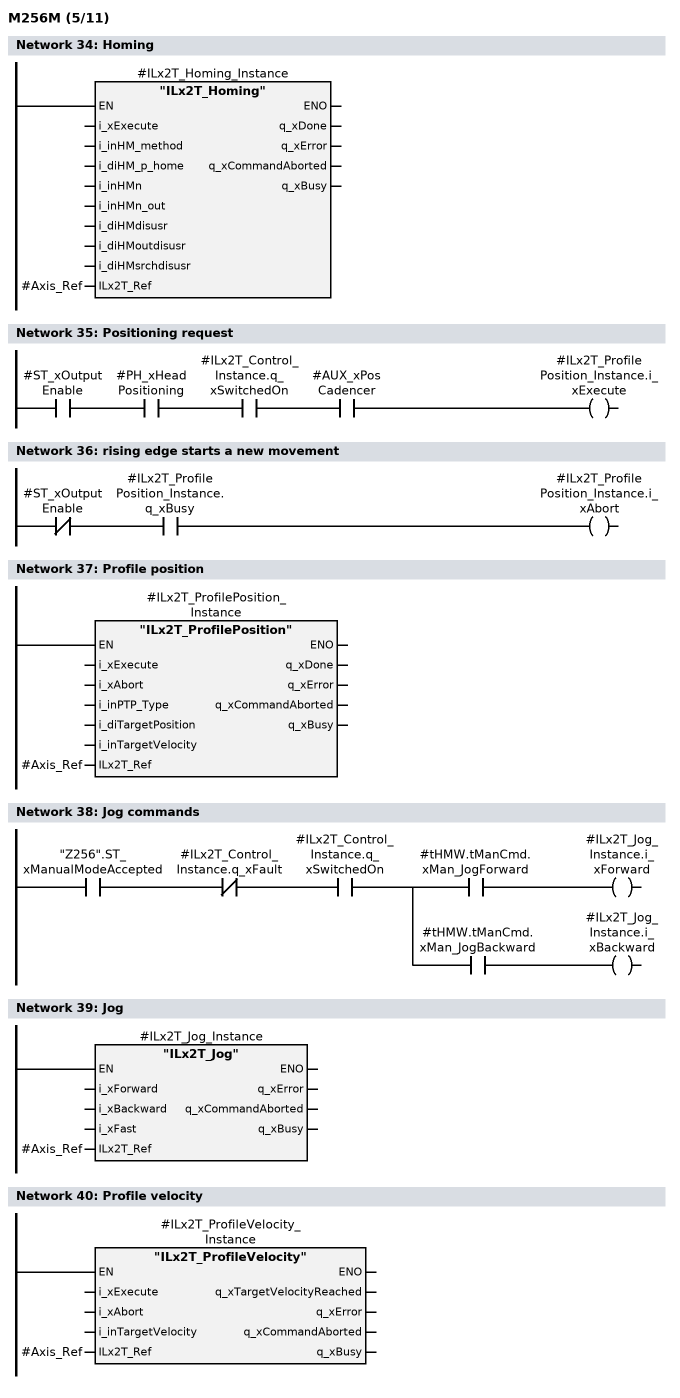
   RUNG wire#powerrail
      #ILx2T_Homing_Instance(i_xExecute :=, i_inHM_method :=, i_diHM_p_home :=, i_inHMn :=, i_inHMn_out :=, i_diHMdisusr :=, i_diHMoutdisusr :=, i_diHMsrchdisusr :=, ILx2T_Ref := #Axis_Ref, q_xDone =>, q_xError =>, q_xCommandAborted =>, q_xBusy =>)
   END_RUNG
   // the same network as SCL:
   #ILx2T_Homing_Instance(ILx2T_Ref := #Axis_Ref);   // "ILx2T_Homing"
END_REGION

REGION Network 35: Positioning request
   RUNG wire#powerrail
      Contact( #ST_xOutputEnable )
      Contact( #PH_xHeadPositioning )
      Contact( #ILx2T_Control_Instance.q_xSwitchedOn )
      Contact( #AUX_xPosCadencer )
      Coil( #ILx2T_ProfilePosition_Instance.i_xExecute )
   END_RUNG
   // the same network as SCL:
   #ILx2T_ProfilePosition_Instance.i_xExecute := #ST_xOutputEnable AND #PH_xHeadPositioning AND #ILx2T_Control_Instance.q_xSwitchedOn AND #AUX_xPosCadencer;
END_REGION

REGION Network 36: rising edge starts a new movement
   RUNG wire#powerrail
      I_Contact( #ST_xOutputEnable )
      Contact( #ILx2T_ProfilePosition_Instance.q_xBusy )
      Coil( #ILx2T_ProfilePosition_Instance.i_xAbort )
   END_RUNG
   // the same network as SCL:
   #ILx2T_ProfilePosition_Instance.i_xAbort := NOT #ST_xOutputEnable AND #ILx2T_ProfilePosition_Instance.q_xBusy;
END_REGION

REGION Network 37: Profile position
   RUNG wire#powerrail
      #ILx2T_ProfilePosition_Instance(i_xExecute :=, i_xAbort :=, i_inPTP_Type :=, i_diTargetPosition :=, i_inTargetVelocity :=, ILx2T_Ref := #Axis_Ref, q_xDone =>, q_xError =>, q_xCommandAborted =>, q_xBusy =>)
   END_RUNG
   // the same network as SCL:
   #ILx2T_ProfilePosition_Instance(ILx2T_Ref := #Axis_Ref);   // "ILx2T_ProfilePosition"
END_REGION

REGION Network 38: Jog commands
   RUNG wire#powerrail
      Contact( "Z256".ST_xManualModeAccepted )
      I_Contact( #ILx2T_Control_Instance.q_xFault )
      Contact( #ILx2T_Control_Instance.q_xSwitchedOn )
      wire#w1
      Contact( #tHMW.tManCmd.xMan_JogForward )
      Coil( #ILx2T_Jog_Instance.i_xForward )
   END_RUNG
   RUNG wire#w1
      Contact( #tHMW.tManCmd.xMan_JogBackward )
      Coil( #ILx2T_Jog_Instance.i_xBackward )
   END_RUNG
   // the same network as SCL:
   #_w1 := "Z256".ST_xManualModeAccepted AND NOT #ILx2T_Control_Instance.q_xFault AND #ILx2T_Control_Instance.q_xSwitchedOn;
   #ILx2T_Jog_Instance.i_xForward := #_w1 AND #tHMW.tManCmd.xMan_JogForward;
   #ILx2T_Jog_Instance.i_xBackward := #_w1 AND #tHMW.tManCmd.xMan_JogBackward;
END_REGION

REGION Network 39: Jog
   RUNG wire#powerrail
      #ILx2T_Jog_Instance(i_xForward :=, i_xBackward :=, i_xFast :=, ILx2T_Ref := #Axis_Ref, q_xError =>, q_xCommandAborted =>, q_xBusy =>)
   END_RUNG
   // the same network as SCL:
   #ILx2T_Jog_Instance(ILx2T_Ref := #Axis_Ref);   // "ILx2T_Jog"
END_REGION

REGION Network 40: Profile velocity
   RUNG wire#powerrail
      #ILx2T_ProfileVelocity_Instance(i_xExecute :=, i_xAbort :=, i_inTargetVelocity :=, ILx2T_Ref := #Axis_Ref, q_xTargetVelocityReached =>, q_xError =>, q_xCommandAborted =>, q_xBusy =>)
   END_RUNG
   // the same network as SCL:
   #ILx2T_ProfileVelocity_Instance(ILx2T_Ref := #Axis_Ref);   // "ILx2T_ProfileVelocity"
END_REGION

REGION Network 41: Head brake release
   // state 3=switch on disabled
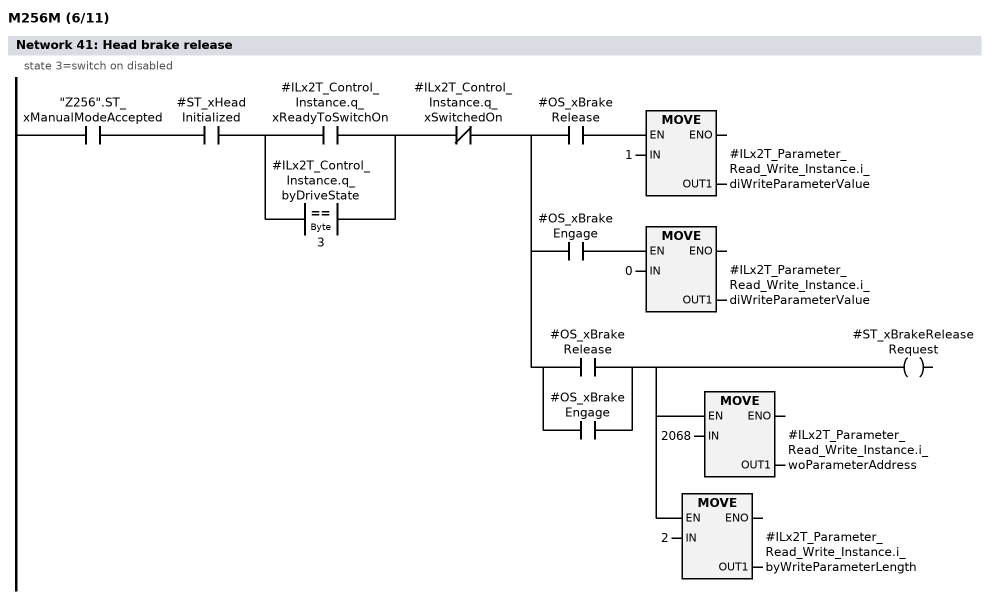
   RUNG wire#powerrail
      Contact( "Z256".ST_xManualModeAccepted )
      Contact( #ST_xHeadInitialized )
      wire#w1
      Contact( #ILx2T_Control_Instance.q_xReadyToSwitchOn )
      wire#w2
      I_Contact( #ILx2T_Control_Instance.q_xSwitchedOn )
      wire#w3
      Contact( #OS_xBrakeRelease )
      Move(in := 1, out1 => #ILx2T_Parameter_Read_Write_Instance.i_diWriteParameterValue)
   END_RUNG
   RUNG wire#w1
      { S7_Templates := "SrcType := Byte" } EQ_Contact(in1 := #ILx2T_Control_Instance.q_byDriveState, in2 := 3)
   END_RUNG wire#w2
   RUNG wire#w3
      Contact( #OS_xBrakeEngage )
      Move(in := 0, out1 => #ILx2T_Parameter_Read_Write_Instance.i_diWriteParameterValue)
   END_RUNG
   RUNG wire#w3
      Contact( #OS_xBrakeRelease )
      wire#w4
      Coil( #ST_xBrakeReleaseRequest )
   END_RUNG
   RUNG wire#w3
      Contact( #OS_xBrakeEngage )
   END_RUNG wire#w4
   RUNG wire#w4
      Move(in := 2068, out1 => #ILx2T_Parameter_Read_Write_Instance.i_woParameterAddress)
   END_RUNG
   RUNG wire#w4
      Move(in := 2, out1 => #ILx2T_Parameter_Read_Write_Instance.i_byWriteParameterLength)
   END_RUNG
   // the same network as SCL:
   #_w1 := "Z256".ST_xManualModeAccepted AND #ST_xHeadInitialized AND (#ILx2T_Control_Instance.q_xReadyToSwitchOn OR (#ILx2T_Control_Instance.q_byDriveState = 3)) AND NOT #ILx2T_Control_Instance.q_xSwitchedOn;
   IF #_w1 AND #OS_xBrakeRelease THEN
       #ILx2T_Parameter_Read_Write_Instance.i_diWriteParameterValue := 1;
   END_IF;
   IF #_w1 AND #OS_xBrakeEngage THEN
       #ILx2T_Parameter_Read_Write_Instance.i_diWriteParameterValue := 0;
   END_IF;
   #ST_xBrakeReleaseRequest := #_w1 AND (#OS_xBrakeRelease OR #OS_xBrakeEngage);
   IF #ST_xBrakeReleaseRequest THEN
       #ILx2T_Parameter_Read_Write_Instance.i_woParameterAddress := 2068;
       #ILx2T_Parameter_Read_Write_Instance.i_byWriteParameterLength := 2;
   END_IF;
END_REGION

REGION Network 42: #### CALCULATE STATUSES ####
END_REGION

REGION Network 43: Read position and speed
   // 5.0 mm / rivoluzione
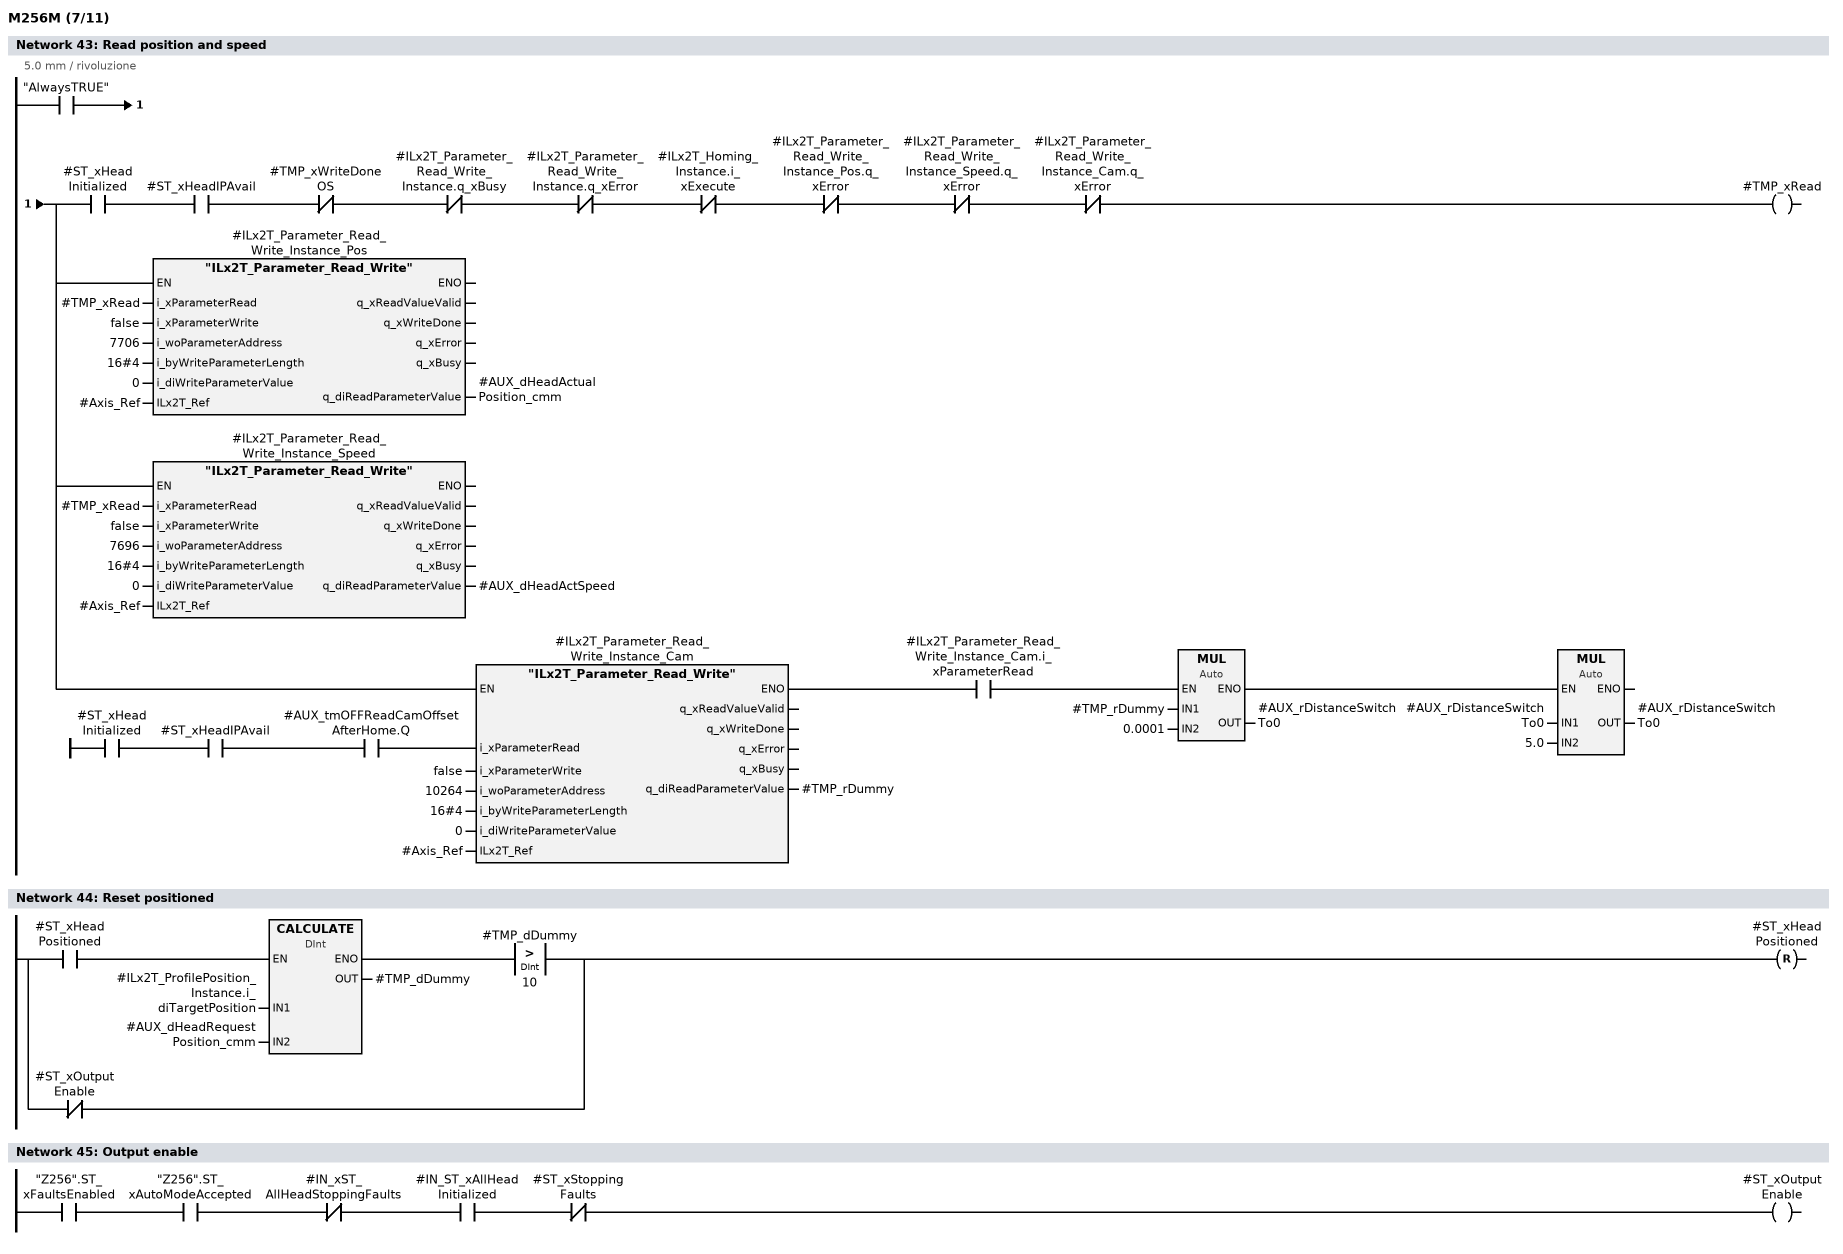
   RUNG wire#powerrail
      Contact( "AlwaysTRUE" )
      wire#w1
      Contact( #ST_xHeadInitialized )
      Contact( #ST_xHeadIPAvail )
      I_Contact( #TMP_xWriteDoneOS )
      I_Contact( #ILx2T_Parameter_Read_Write_Instance.q_xBusy )
      I_Contact( #ILx2T_Parameter_Read_Write_Instance.q_xError )
      I_Contact( #ILx2T_Homing_Instance.i_xExecute )
      I_Contact( #ILx2T_Parameter_Read_Write_Instance_Pos.q_xError )
      I_Contact( #ILx2T_Parameter_Read_Write_Instance_Speed.q_xError )
      I_Contact( #ILx2T_Parameter_Read_Write_Instance_Cam.q_xError )
      Coil( #TMP_xRead )
   END_RUNG
   RUNG wire#w1
      #ILx2T_Parameter_Read_Write_Instance_Pos(i_xParameterRead := #TMP_xRead, i_xParameterWrite := false, i_woParameterAddress := 7706, i_byWriteParameterLength := 16#4, i_diWriteParameterValue := 0, ILx2T_Ref := #Axis_Ref, q_xReadValueValid =>, q_xWriteDone =>, q_xError =>, q_xBusy =>, q_diReadParameterValue => #AUX_dHeadActualPosition_cmm)
   END_RUNG
   RUNG wire#w1
      #ILx2T_Parameter_Read_Write_Instance_Speed(i_xParameterRead := #TMP_xRead, i_xParameterWrite := false, i_woParameterAddress := 7696, i_byWriteParameterLength := 16#4, i_diWriteParameterValue := 0, ILx2T_Ref := #Axis_Ref, q_xReadValueValid =>, q_xWriteDone =>, q_xError =>, q_xBusy =>, q_diReadParameterValue => #AUX_dHeadActSpeed)
   END_RUNG
   RUNG wire#w1
      #ILx2T_Parameter_Read_Write_Instance_Cam(i_xParameterRead := wire#w2, i_xParameterWrite := false, i_woParameterAddress := 10264, i_byWriteParameterLength := 16#4, i_diWriteParameterValue := 0, ILx2T_Ref := #Axis_Ref, q_xReadValueValid =>, q_xWriteDone =>, q_xError =>, q_xBusy =>, q_diReadParameterValue => #TMP_rDummy)
      Contact( #ILx2T_Parameter_Read_Write_Instance_Cam.i_xParameterRead )
      Mul(in1 := #TMP_rDummy, in2 := 0.0001, out => #AUX_rDistanceSwitchTo0)
      Mul(in1 := #AUX_rDistanceSwitchTo0, in2 := 5.0, out => #AUX_rDistanceSwitchTo0)
   END_RUNG
   RUNG wire#powerrail
      Contact( #ST_xHeadInitialized )
      Contact( #ST_xHeadIPAvail )
      Contact( #AUX_tmOFFReadCamOffsetAfterHome.Q )
   END_RUNG wire#w2
   // the same network as SCL:
   #TMP_xRead := "AlwaysTRUE" AND #ST_xHeadInitialized AND #ST_xHeadIPAvail AND NOT #TMP_xWriteDoneOS AND NOT #ILx2T_Parameter_Read_Write_Instance.q_xBusy AND NOT #ILx2T_Parameter_Read_Write_Instance.q_xError AND NOT #ILx2T_Homing_Instance.i_xExecute AND NOT #ILx2T_Parameter_Read_Write_Instance_Pos.q_xError AND NOT #ILx2T_Parameter_Read_Write_Instance_Speed.q_xError AND NOT #ILx2T_Parameter_Read_Write_Instance_Cam.q_xError;
   #_w1 := "AlwaysTRUE";
   IF #_w1 THEN
       #ILx2T_Parameter_Read_Write_Instance_Pos(i_xParameterRead := #TMP_xRead,   // "ILx2T_Parameter_Read_Write"
                               i_xParameterWrite := false,
                               i_woParameterAddress := 7706,
                               i_byWriteParameterLength := 16#4,
                               i_diWriteParameterValue := 0,
                               ILx2T_Ref := #Axis_Ref,
                               q_diReadParameterValue => #AUX_dHeadActualPosition_cmm);
       #ILx2T_Parameter_Read_Write_Instance_Speed(i_xParameterRead := #TMP_xRead,   // "ILx2T_Parameter_Read_Write"
                               i_xParameterWrite := false,
                               i_woParameterAddress := 7696,
                               i_byWriteParameterLength := 16#4,
                               i_diWriteParameterValue := 0,
                               ILx2T_Ref := #Axis_Ref,
                               q_diReadParameterValue => #AUX_dHeadActSpeed);
   END_IF;
   #ILx2T_Parameter_Read_Write_Instance_Cam(EN := #_w1,   // "ILx2T_Parameter_Read_Write"
                           i_xParameterRead := #ST_xHeadInitialized AND #ST_xHeadIPAvail AND #AUX_tmOFFReadCamOffsetAfterHome.Q,
                           i_xParameterWrite := false,
                           i_woParameterAddress := 10264,
                           i_byWriteParameterLength := 16#4,
                           i_diWriteParameterValue := 0,
                           ILx2T_Ref := #Axis_Ref,
                           q_diReadParameterValue => #TMP_rDummy,
                           ENO => #_w2);
   IF #_w2 AND #ILx2T_Parameter_Read_Write_Instance_Cam.i_xParameterRead THEN
       #AUX_rDistanceSwitchTo0 := #TMP_rDummy * 0.0001;
       #AUX_rDistanceSwitchTo0 := #AUX_rDistanceSwitchTo0 * 5.0;
   END_IF;
END_REGION

REGION Network 44: Reset positioned
   RUNG wire#powerrail
      Contact( #ST_xHeadPositioned )
      { S7_Templates := "SrcType := DInt"; S7_Expression := "ABS(IN2-IN1)" } Calculate(in1 := #ILx2T_ProfilePosition_Instance.i_diTargetPosition, in2 := #AUX_dHeadRequestPosition_cmm, out => #TMP_dDummy)
      { S7_Templates := "SrcType := DInt" } GT_Contact(in1 := #TMP_dDummy, in2 := 10)
      wire#w1
      R_Coil( #ST_xHeadPositioned )
   END_RUNG
   RUNG wire#powerrail
      I_Contact( #ST_xOutputEnable )
   END_RUNG wire#w1
   // the same network as SCL:
   IF #ST_xHeadPositioned THEN
       #TMP_dDummy := ABS(#AUX_dHeadRequestPosition_cmm-#ILx2T_ProfilePosition_Instance.i_diTargetPosition);
   END_IF;
   IF (#ST_xHeadPositioned AND (#TMP_dDummy > 10)) OR NOT #ST_xOutputEnable THEN
       #ST_xHeadPositioned := FALSE;
   END_IF;
END_REGION

REGION Network 45: Output enable
   RUNG wire#powerrail
      Contact( "Z256".ST_xFaultsEnabled )
      Contact( "Z256".ST_xAutoModeAccepted )
      I_Contact( #IN_xST_AllHeadStoppingFaults )
      Contact( #IN_ST_xAllHeadInitialized )
      I_Contact( #ST_xStoppingFaults )
      Coil( #ST_xOutputEnable )
   END_RUNG
   // the same network as SCL:
   #ST_xOutputEnable := "Z256".ST_xFaultsEnabled AND "Z256".ST_xAutoModeAccepted AND NOT #IN_xST_AllHeadStoppingFaults AND #IN_ST_xAllHeadInitialized AND NOT #ST_xStoppingFaults;
END_REGION

REGION Network 46: Head #x in movement
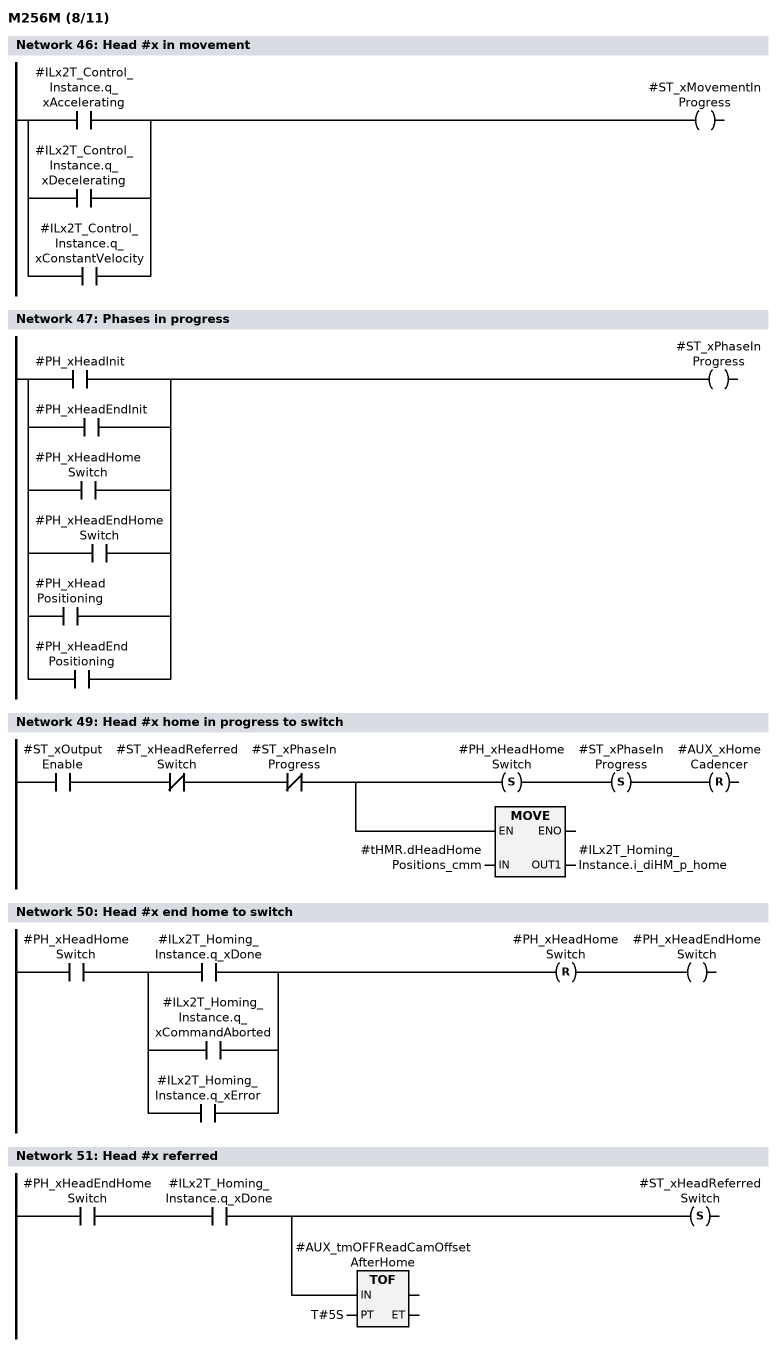
   RUNG wire#powerrail
      Contact( #ILx2T_Control_Instance.q_xAccelerating )
      wire#w1
      Coil( #ST_xMovementInProgress )
   END_RUNG
   RUNG wire#powerrail
      Contact( #ILx2T_Control_Instance.q_xDecelerating )
   END_RUNG wire#w1
   RUNG wire#powerrail
      Contact( #ILx2T_Control_Instance.q_xConstantVelocity )
   END_RUNG wire#w1
   // the same network as SCL:
   #ST_xMovementInProgress := #ILx2T_Control_Instance.q_xAccelerating OR #ILx2T_Control_Instance.q_xDecelerating OR #ILx2T_Control_Instance.q_xConstantVelocity;
END_REGION

REGION Network 47: Phases in progress
   RUNG wire#powerrail
      Contact( #PH_xHeadInit )
      wire#w1
      Coil( #ST_xPhaseInProgress )
   END_RUNG
   RUNG wire#powerrail
      Contact( #PH_xHeadEndInit )
   END_RUNG wire#w1
   RUNG wire#powerrail
      Contact( #PH_xHeadHomeSwitch )
   END_RUNG wire#w1
   RUNG wire#powerrail
      Contact( #PH_xHeadEndHomeSwitch )
   END_RUNG wire#w1
   RUNG wire#powerrail
      Contact( #PH_xHeadPositioning )
   END_RUNG wire#w1
   RUNG wire#powerrail
      Contact( #PH_xHeadEndPositioning )
   END_RUNG wire#w1
   // the same network as SCL:
   #ST_xPhaseInProgress := #PH_xHeadInit OR #PH_xHeadEndInit OR #PH_xHeadHomeSwitch OR #PH_xHeadEndHomeSwitch OR #PH_xHeadPositioning OR #PH_xHeadEndPositioning;
END_REGION

REGION Network 48: #### CALCULATE PHASES ####
END_REGION

REGION Network 49: Head #x home in progress to switch
   RUNG wire#powerrail
      Contact( #ST_xOutputEnable )
      I_Contact( #ST_xHeadReferredSwitch )
      I_Contact( #ST_xPhaseInProgress )
      wire#w1
      S_Coil( #PH_xHeadHomeSwitch )
      S_Coil( #ST_xPhaseInProgress )
      R_Coil( #AUX_xHomeCadencer )
   END_RUNG
   RUNG wire#w1
      Move(in := #tHMR.dHeadHomePositions_cmm, out1 => #ILx2T_Homing_Instance.i_diHM_p_home)
   END_RUNG
   // the same network as SCL:
   IF #ST_xOutputEnable AND NOT #ST_xHeadReferredSwitch AND NOT #ST_xPhaseInProgress THEN
       #PH_xHeadHomeSwitch := TRUE;
   END_IF;
   #_w1 := #ST_xOutputEnable AND NOT #ST_xHeadReferredSwitch AND NOT #ST_xPhaseInProgress;
   IF #_w1 THEN
       #ST_xPhaseInProgress := TRUE;
       #AUX_xHomeCadencer := FALSE;
       #ILx2T_Homing_Instance.i_diHM_p_home := #tHMR.dHeadHomePositions_cmm;
   END_IF;
END_REGION

REGION Network 50: Head #x end home to switch
   RUNG wire#powerrail
      Contact( #PH_xHeadHomeSwitch )
      wire#w1
      Contact( #ILx2T_Homing_Instance.q_xDone )
      wire#w2
      R_Coil( #PH_xHeadHomeSwitch )
      Coil( #PH_xHeadEndHomeSwitch )
   END_RUNG
   RUNG wire#w1
      Contact( #ILx2T_Homing_Instance.q_xCommandAborted )
   END_RUNG wire#w2
   RUNG wire#w1
      Contact( #ILx2T_Homing_Instance.q_xError )
   END_RUNG wire#w2
   // the same network as SCL:
   #_w1 := #PH_xHeadHomeSwitch AND (#ILx2T_Homing_Instance.q_xDone OR #ILx2T_Homing_Instance.q_xCommandAborted OR #ILx2T_Homing_Instance.q_xError);
   IF #_w1 THEN #PH_xHeadHomeSwitch := FALSE; END_IF;
   #PH_xHeadEndHomeSwitch := #_w1;
END_REGION

REGION Network 51: Head #x referred
   #_w1 := #PH_xHeadEndHomeSwitch AND #ILx2T_Homing_Instance.q_xDone;
   IF #_w1 THEN #ST_xHeadReferredSwitch := TRUE; END_IF;
   #AUX_tmOFFReadCamOffsetAfterHome.TOF(IN := #_w1, PT := T#5S);
END_REGION

REGION Network 52: Wait positioning after home
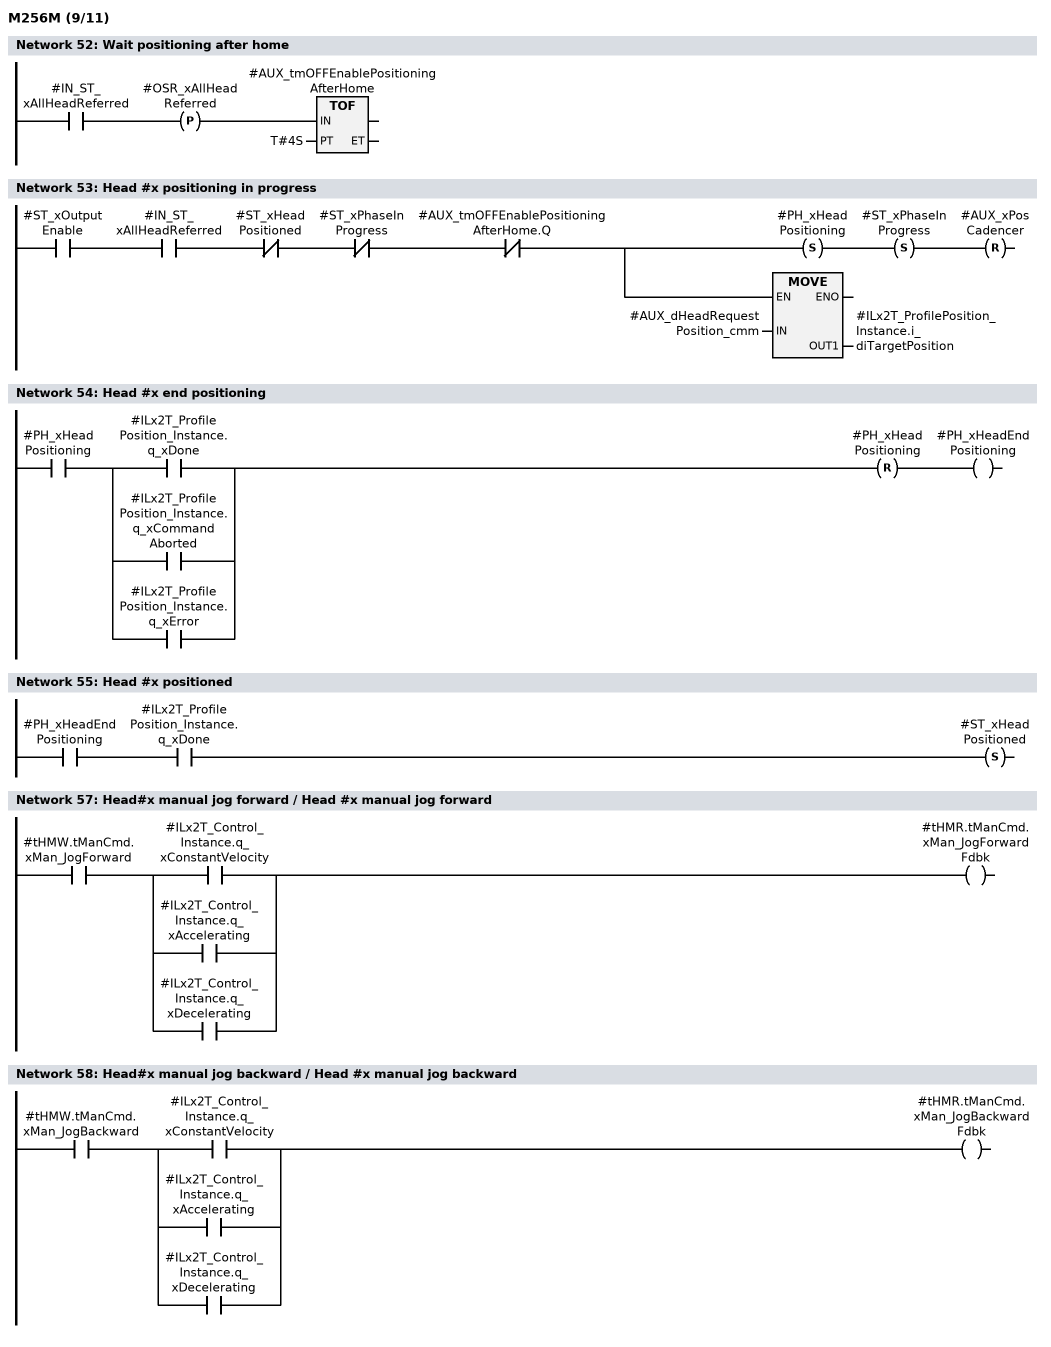
   #_w1 := #IN_ST_xAllHeadReferred AND NOT #OSR_xAllHeadReferred;   // rising edge
   #OSR_xAllHeadReferred := #IN_ST_xAllHeadReferred;
   #AUX_tmOFFEnablePositioningAfterHome.TOF(IN := #_w1, PT := T#4S);
END_REGION

REGION Network 53: Head #x positioning in progress
   RUNG wire#powerrail
      Contact( #ST_xOutputEnable )
      Contact( #IN_ST_xAllHeadReferred )
      I_Contact( #ST_xHeadPositioned )
      I_Contact( #ST_xPhaseInProgress )
      I_Contact( #AUX_tmOFFEnablePositioningAfterHome.Q )
      wire#w1
      S_Coil( #PH_xHeadPositioning )
      S_Coil( #ST_xPhaseInProgress )
      R_Coil( #AUX_xPosCadencer )
   END_RUNG
   RUNG wire#w1
      Move(in := #AUX_dHeadRequestPosition_cmm, out1 => #ILx2T_ProfilePosition_Instance.i_diTargetPosition)
   END_RUNG
   // the same network as SCL:
   IF #ST_xOutputEnable AND #IN_ST_xAllHeadReferred AND NOT #ST_xHeadPositioned AND NOT #ST_xPhaseInProgress AND NOT #AUX_tmOFFEnablePositioningAfterHome.Q THEN
       #PH_xHeadPositioning := TRUE;
   END_IF;
   #_w1 := #ST_xOutputEnable AND #IN_ST_xAllHeadReferred AND NOT #ST_xHeadPositioned AND NOT #ST_xPhaseInProgress AND NOT #AUX_tmOFFEnablePositioningAfterHome.Q;
   IF #_w1 THEN
       #ST_xPhaseInProgress := TRUE;
       #AUX_xPosCadencer := FALSE;
       #ILx2T_ProfilePosition_Instance.i_diTargetPosition := #AUX_dHeadRequestPosition_cmm;
   END_IF;
END_REGION

REGION Network 54: Head #x end positioning
   RUNG wire#powerrail
      Contact( #PH_xHeadPositioning )
      wire#w1
      Contact( #ILx2T_ProfilePosition_Instance.q_xDone )
      wire#w2
      R_Coil( #PH_xHeadPositioning )
      Coil( #PH_xHeadEndPositioning )
   END_RUNG
   RUNG wire#w1
      Contact( #ILx2T_ProfilePosition_Instance.q_xCommandAborted )
   END_RUNG wire#w2
   RUNG wire#w1
      Contact( #ILx2T_ProfilePosition_Instance.q_xError )
   END_RUNG wire#w2
   // the same network as SCL:
   #_w1 := #PH_xHeadPositioning AND (#ILx2T_ProfilePosition_Instance.q_xDone OR #ILx2T_ProfilePosition_Instance.q_xCommandAborted OR #ILx2T_ProfilePosition_Instance.q_xError);
   IF #_w1 THEN #PH_xHeadPositioning := FALSE; END_IF;
   #PH_xHeadEndPositioning := #_w1;
END_REGION

REGION Network 55: Head #x positioned
   RUNG wire#powerrail
      Contact( #PH_xHeadEndPositioning )
      Contact( #ILx2T_ProfilePosition_Instance.q_xDone )
      S_Coil( #ST_xHeadPositioned )
   END_RUNG
   // the same network as SCL:
   IF #PH_xHeadEndPositioning AND #ILx2T_ProfilePosition_Instance.q_xDone THEN
       #ST_xHeadPositioned := TRUE;
   END_IF;
END_REGION

REGION Network 56: #### HMI STATUSES ####
END_REGION

REGION Network 57: Head#x manual jog forward / Head #x manual jog forward
   RUNG wire#powerrail
      Contact( #tHMW.tManCmd.xMan_JogForward )
      wire#w1
      Contact( #ILx2T_Control_Instance.q_xConstantVelocity )
      wire#w2
      Coil( #tHMR.tManCmd.xMan_JogForwardFdbk )
   END_RUNG
   RUNG wire#w1
      Contact( #ILx2T_Control_Instance.q_xAccelerating )
   END_RUNG wire#w2
   RUNG wire#w1
      Contact( #ILx2T_Control_Instance.q_xDecelerating )
   END_RUNG wire#w2
   // the same network as SCL:
   #tHMR.tManCmd.xMan_JogForwardFdbk := #tHMW.tManCmd.xMan_JogForward AND (#ILx2T_Control_Instance.q_xConstantVelocity OR #ILx2T_Control_Instance.q_xAccelerating OR #ILx2T_Control_Instance.q_xDecelerating);
END_REGION

REGION Network 58: Head#x manual jog backward / Head #x manual jog backward
   RUNG wire#powerrail
      Contact( #tHMW.tManCmd.xMan_JogBackward )
      wire#w1
      Contact( #ILx2T_Control_Instance.q_xConstantVelocity )
      wire#w2
      Coil( #tHMR.tManCmd.xMan_JogBackwardFdbk )
   END_RUNG
   RUNG wire#w1
      Contact( #ILx2T_Control_Instance.q_xAccelerating )
   END_RUNG wire#w2
   RUNG wire#w1
      Contact( #ILx2T_Control_Instance.q_xDecelerating )
   END_RUNG wire#w2
   // the same network as SCL:
   #tHMR.tManCmd.xMan_JogBackwardFdbk := #tHMW.tManCmd.xMan_JogBackward AND (#ILx2T_Control_Instance.q_xConstantVelocity OR #ILx2T_Control_Instance.q_xAccelerating OR #ILx2T_Control_Instance.q_xDecelerating);
END_REGION

REGION Network 59: Head status
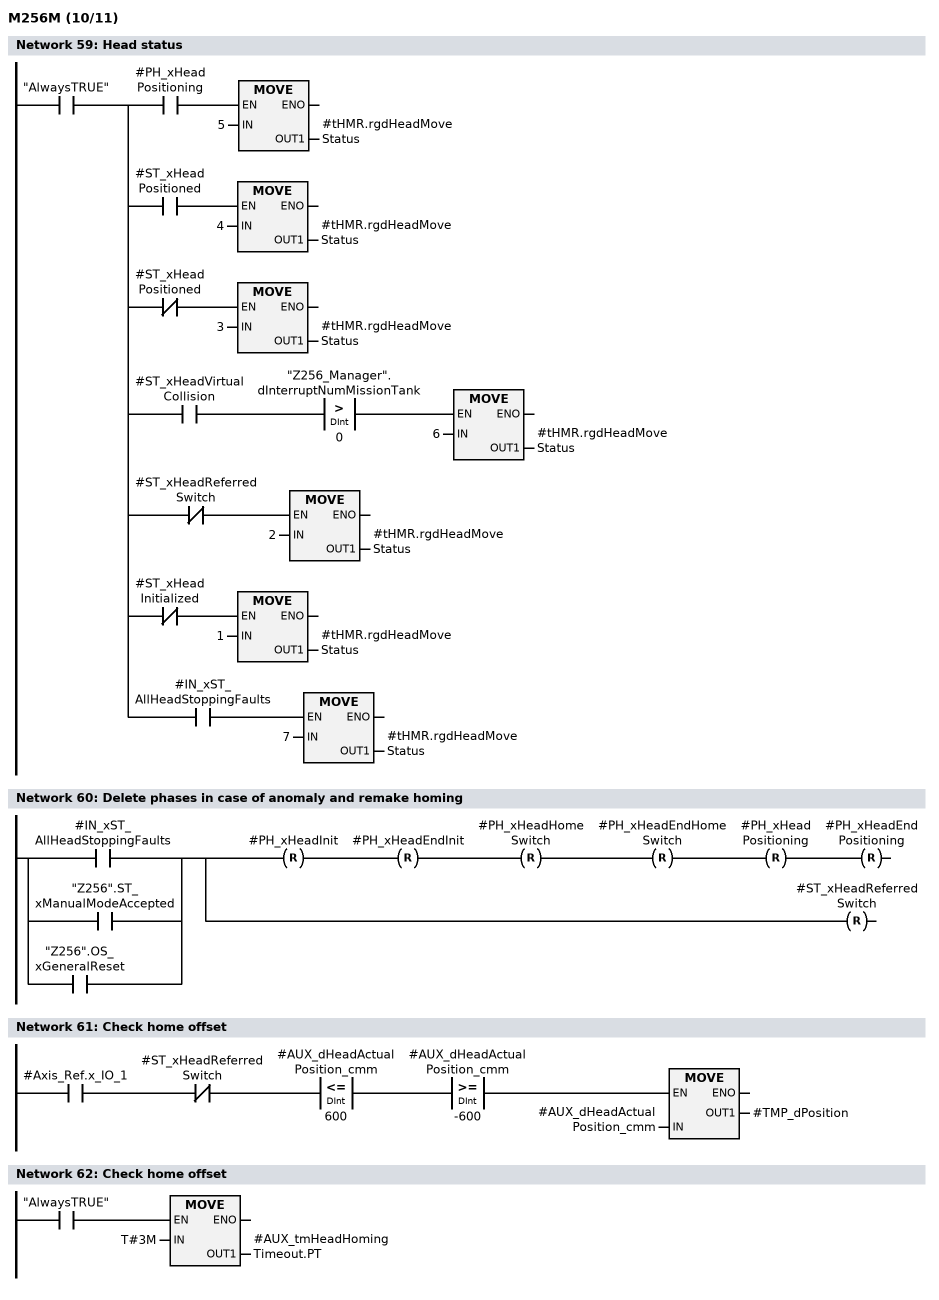
   RUNG wire#powerrail
      Contact( "AlwaysTRUE" )
      wire#w1
      Contact( #PH_xHeadPositioning )
      Move(in := 5, out1 => #tHMR.rgdHeadMoveStatus)
   END_RUNG
   RUNG wire#w1
      Contact( #ST_xHeadPositioned )
      Move(in := 4, out1 => #tHMR.rgdHeadMoveStatus)
   END_RUNG
   RUNG wire#w1
      I_Contact( #ST_xHeadPositioned )
      Move(in := 3, out1 => #tHMR.rgdHeadMoveStatus)
   END_RUNG
   RUNG wire#w1
      Contact( #ST_xHeadVirtualCollision )
      { S7_Templates := "SrcType := DInt" } GT_Contact(in1 := "Z256_Manager".dInterruptNumMissionTank, in2 := 0)
      Move(in := 6, out1 => #tHMR.rgdHeadMoveStatus)
   END_RUNG
   RUNG wire#w1
      I_Contact( #ST_xHeadReferredSwitch )
      Move(in := 2, out1 => #tHMR.rgdHeadMoveStatus)
   END_RUNG
   RUNG wire#w1
      I_Contact( #ST_xHeadInitialized )
      Move(in := 1, out1 => #tHMR.rgdHeadMoveStatus)
   END_RUNG
   RUNG wire#w1
      Contact( #IN_xST_AllHeadStoppingFaults )
      Move(in := 7, out1 => #tHMR.rgdHeadMoveStatus)
   END_RUNG
   // the same network as SCL:
   IF "AlwaysTRUE" AND #PH_xHeadPositioning THEN #tHMR.rgdHeadMoveStatus := 5; END_IF;
   IF "AlwaysTRUE" AND #ST_xHeadPositioned THEN #tHMR.rgdHeadMoveStatus := 4; END_IF;
   IF "AlwaysTRUE" AND NOT #ST_xHeadPositioned THEN #tHMR.rgdHeadMoveStatus := 3; END_IF;
   IF "AlwaysTRUE" AND #ST_xHeadVirtualCollision AND ("Z256_Manager".dInterruptNumMissionTank > 0) THEN
       #tHMR.rgdHeadMoveStatus := 6;
   END_IF;
   IF "AlwaysTRUE" AND NOT #ST_xHeadReferredSwitch THEN #tHMR.rgdHeadMoveStatus := 2; END_IF;
   IF "AlwaysTRUE" AND NOT #ST_xHeadInitialized THEN #tHMR.rgdHeadMoveStatus := 1; END_IF;
   IF "AlwaysTRUE" AND #IN_xST_AllHeadStoppingFaults THEN #tHMR.rgdHeadMoveStatus := 7; END_IF;
END_REGION

REGION Network 60: Delete phases in case of anomaly and remake homing
   RUNG wire#powerrail
      Contact( #IN_xST_AllHeadStoppingFaults )
      wire#w1
      R_Coil( #PH_xHeadInit )
      R_Coil( #PH_xHeadEndInit )
      R_Coil( #PH_xHeadHomeSwitch )
      R_Coil( #PH_xHeadEndHomeSwitch )
      R_Coil( #PH_xHeadPositioning )
      R_Coil( #PH_xHeadEndPositioning )
   END_RUNG
   RUNG wire#powerrail
      Contact( "Z256".ST_xManualModeAccepted )
   END_RUNG wire#w1
   RUNG wire#powerrail
      Contact( "Z256".OS_xGeneralReset )
   END_RUNG wire#w1
   RUNG wire#w1
      R_Coil( #ST_xHeadReferredSwitch )
   END_RUNG
   // the same network as SCL:
   IF #IN_xST_AllHeadStoppingFaults OR "Z256".ST_xManualModeAccepted OR "Z256".OS_xGeneralReset THEN
       #PH_xHeadInit := FALSE;
       #PH_xHeadEndInit := FALSE;
       #PH_xHeadHomeSwitch := FALSE;
       #PH_xHeadEndHomeSwitch := FALSE;
       #PH_xHeadPositioning := FALSE;
       #PH_xHeadEndPositioning := FALSE;
       #ST_xHeadReferredSwitch := FALSE;
   END_IF;
END_REGION

REGION Network 61: Check home offset
   RUNG wire#powerrail
      Contact( #Axis_Ref.x_IO_1 )
      I_Contact( #ST_xHeadReferredSwitch )
      { S7_Templates := "SrcType := DInt" } LE_Contact(in1 := #AUX_dHeadActualPosition_cmm, in2 := 600)
      { S7_Templates := "SrcType := DInt" } GE_Contact(in1 := #AUX_dHeadActualPosition_cmm, in2 := -600)
      Move(in := #AUX_dHeadActualPosition_cmm, out1 => #TMP_dPosition)
   END_RUNG
   // the same network as SCL:
   IF #Axis_Ref.x_IO_1 AND NOT #ST_xHeadReferredSwitch AND (#AUX_dHeadActualPosition_cmm <= 600) AND (#AUX_dHeadActualPosition_cmm >= (-600)) THEN
       #TMP_dPosition := #AUX_dHeadActualPosition_cmm;
   END_IF;
END_REGION

REGION Network 62: Check home offset
   RUNG wire#powerrail
      Contact( "AlwaysTRUE" )
      Move(in := T#3M, out1 => #AUX_tmHeadHomingTimeout.PT)
   END_RUNG
   // the same network as SCL:
   IF "AlwaysTRUE" THEN #AUX_tmHeadHomingTimeout.PT := T#3M; END_IF;
END_REGION

REGION Network 63: Head position
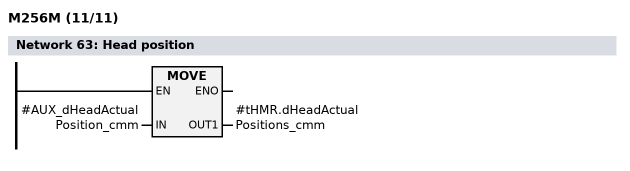
   RUNG wire#powerrail
      Move(in := #AUX_dHeadActualPosition_cmm, out1 => #tHMR.dHeadActualPositions_cmm)
   END_RUNG
   // the same network as SCL:
   #tHMR.dHeadActualPositions_cmm := #AUX_dHeadActualPosition_cmm;
END_REGION
END_FUNCTION_BLOCK

FUNCTION "M256M_SbrCalibrateBridgeOffset" : Void   // FC1, SCL
{ S7_Optimized_Access := 'TRUE' }
VERSION : 0.1
   VAR_IN_OUT
      io_ST_xHeadReferredSwitch : Array[0.."CONST_dNumberOfHeadsCycle"] of Bool;
   END_VAR
   VAR_TEMP
      TMP_dIndex : DInt;
   END_VAR
BEGIN
   ////--------------------------------------------------------------------------------------------------------------------
   //   Copyright (c)  Bottero Spa
   //--------------------------------------------------------------
   //   Routine: CalibratePosition                 
   //       Author: Alberto Cigliutti
   //   Created: <Date>
   //--------------------------------------------------------------
   //   Description: This function will calibrate the bridge offset                
   //
   //   History:
   //
   ////--------------------------------------------------------------------------------------------------------------------

   FOR #TMP_dIndex := 0 TO "CONST_dNumberOfHeadsCycle" DO

       //This function will move the bridge of the requested offset
       //Positive offset all the head move to opposite operatore side
       //Negative offset all the head move to operator side
       //  IF NOT PLANT_CONSTANTS.CONST_RGXHOMESIDE[TMP_dIndex] THEN
       //Operator side
       //Sum the value
       //      M256M_HMR.rgdHeadHomePositions_cmm[TMP_dIndex]  := M256M_HMR.rgdHeadHomePositions_cmm[TMP_dIndex] + M256M_HMW.dMoveBridgeOffset_cmm;
       //  ELSE
       //Opposite operator side
       "M256_Manag_IDB".M256M_IDB[#TMP_dIndex].tHMR.dHeadHomePositions_cmm := "M256_Manag_IDB".M256M_IDB[#TMP_dIndex].tHMR.dHeadHomePositions_cmm - "Z256_hmi".tHMW.dMoveBridgeOffset_cmm;
       //  END_IF;

   END_FOR;

   //Force the heads homing
   FOR #TMP_dIndex := 0 TO "CONST_dNumberOfHeadsCycle" DO
       #io_ST_xHeadReferredSwitch[#TMP_dIndex] := 0;
   END_FOR;
   "Z256_hmi".tHMW.dMoveBridgeOffset_cmm := 0;
END_FUNCTION

FUNCTION "Z256_Logic" : Void   // FC2, LAD
{ S7_Optimized_Access := 'TRUE' }
VERSION : 0.1
   VAR_TEMP
      TMP_iIndex : Int;
      TMP_xDummy : Bool;
      TMP_xCarriageOverload : Bool;
   END_VAR
   VAR_TEMP   // added for the SCL form of the ladder/FBD networks
      _w1 : Bool;
   END_VAR
BEGIN

REGION Network 1: ##### CONSTANTS #####
END_REGION

REGION Network 2: ##### MATCH #####
END_REGION

REGION Network 3: Power alimentation present delayed
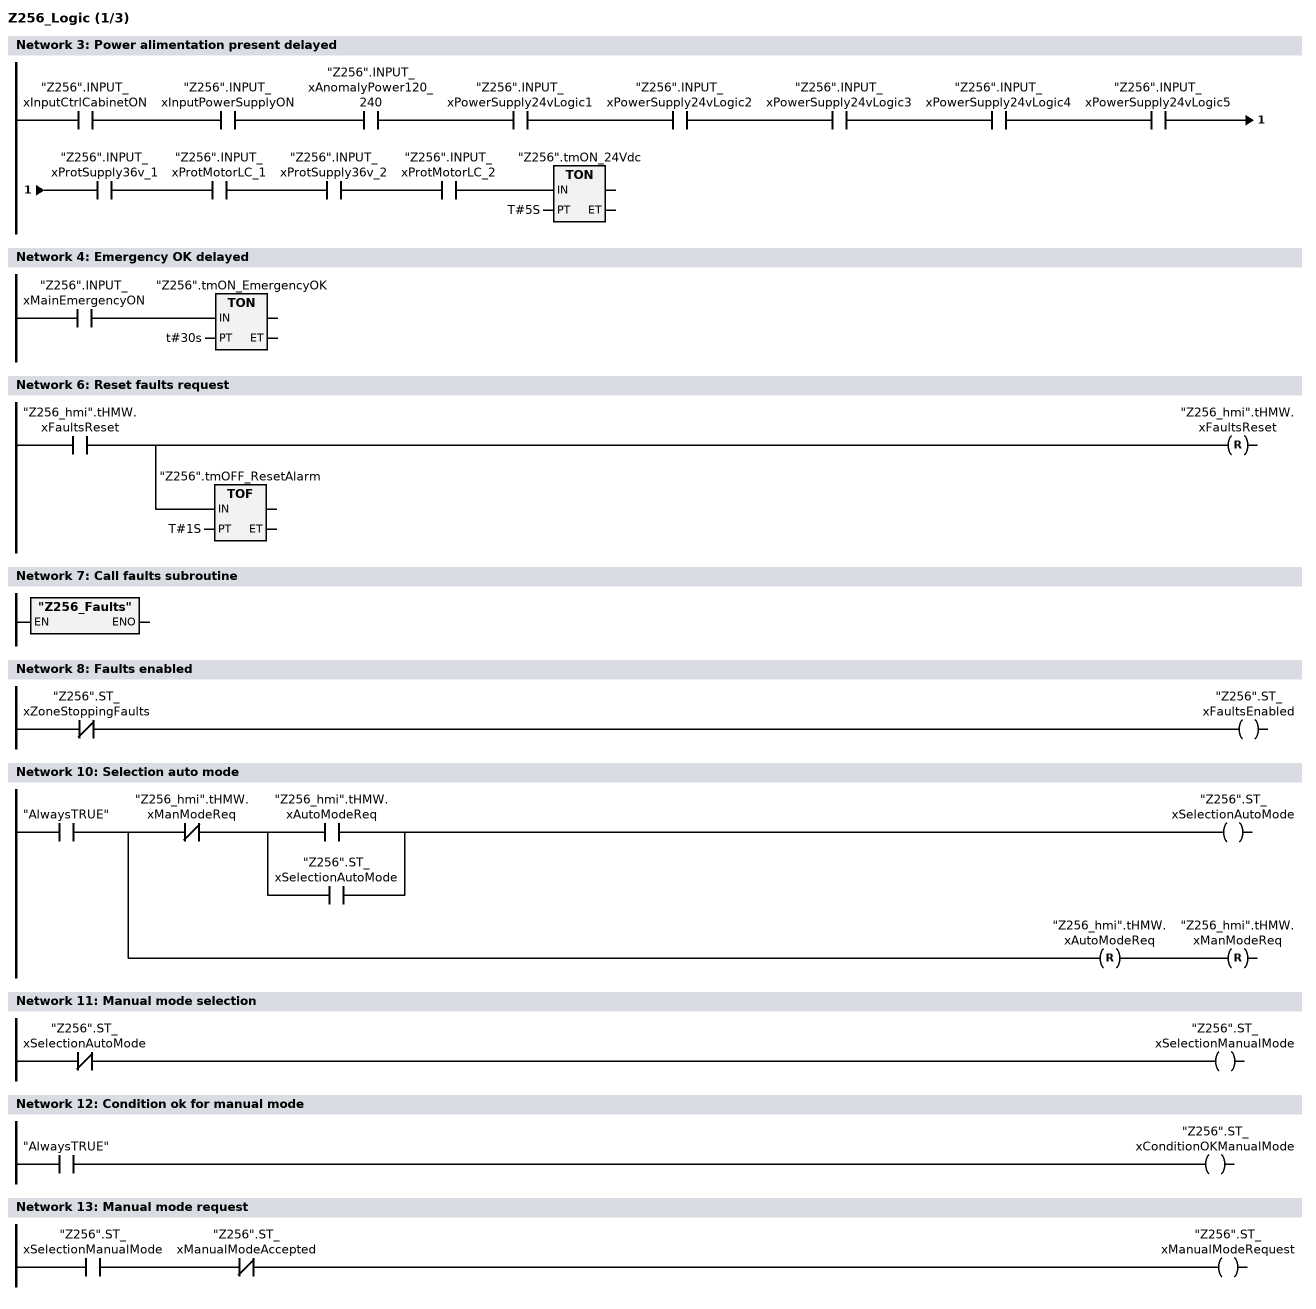
   "Z256".tmON_24Vdc.TON(IN := "Z256".INPUT_xInputCtrlCabinetON AND "Z256".INPUT_xInputPowerSupplyON AND "Z256".INPUT_xAnomalyPower120_240 AND "Z256".INPUT_xPowerSupply24vLogic1 AND "Z256".INPUT_xPowerSupply24vLogic2 AND "Z256".INPUT_xPowerSupply24vLogic3 AND "Z256".INPUT_xPowerSupply24vLogic4 AND "Z256".INPUT_xPowerSupply24vLogic5 AND "Z256".INPUT_xProtSupply36v_1 AND "Z256".INPUT_xProtMotorLC_1 AND "Z256".INPUT_xProtSupply36v_2 AND "Z256".INPUT_xProtMotorLC_2,
                         PT := T#5S);
END_REGION

REGION Network 4: Emergency OK delayed
   "Z256".tmON_EmergencyOK.TON(IN := "Z256".INPUT_xMainEmergencyON, PT := t#30s);
END_REGION

REGION Network 5: ##### FAULTS #####
END_REGION

REGION Network 6: Reset faults request
   #_w1 := "Z256_hmi".tHMW.xFaultsReset;
   IF #_w1 THEN "Z256_hmi".tHMW.xFaultsReset := FALSE; END_IF;
   "Z256".tmOFF_ResetAlarm.TOF(IN := #_w1, PT := T#1S);
END_REGION

REGION Network 7: Call faults subroutine
   RUNG wire#powerrail
      "Z256_Faults"()
   END_RUNG
   // the same network as SCL:
   "Z256_Faults"();
END_REGION

REGION Network 8: Faults enabled
   RUNG wire#powerrail
      I_Contact( "Z256".ST_xZoneStoppingFaults )
      Coil( "Z256".ST_xFaultsEnabled )
   END_RUNG
   // the same network as SCL:
   "Z256".ST_xFaultsEnabled := NOT "Z256".ST_xZoneStoppingFaults;
END_REGION

REGION Network 9: ##### MODE #####
END_REGION

REGION Network 10: Selection auto mode
   RUNG wire#powerrail
      Contact( "AlwaysTRUE" )
      wire#w1
      I_Contact( "Z256_hmi".tHMW.xManModeReq )
      wire#w2
      Contact( "Z256_hmi".tHMW.xAutoModeReq )
      wire#w3
      Coil( "Z256".ST_xSelectionAutoMode )
   END_RUNG
   RUNG wire#w2
      Contact( "Z256".ST_xSelectionAutoMode )
   END_RUNG wire#w3
   RUNG wire#w1
      R_Coil( "Z256_hmi".tHMW.xAutoModeReq )
      R_Coil( "Z256_hmi".tHMW.xManModeReq )
   END_RUNG
   // the same network as SCL:
   "Z256".ST_xSelectionAutoMode := "AlwaysTRUE" AND NOT "Z256_hmi".tHMW.xManModeReq AND ("Z256_hmi".tHMW.xAutoModeReq OR "Z256".ST_xSelectionAutoMode);
   IF "AlwaysTRUE" THEN
       "Z256_hmi".tHMW.xAutoModeReq := FALSE;
       "Z256_hmi".tHMW.xManModeReq := FALSE;
   END_IF;
END_REGION

REGION Network 11: Manual mode selection
   RUNG wire#powerrail
      I_Contact( "Z256".ST_xSelectionAutoMode )
      Coil( "Z256".ST_xSelectionManualMode )
   END_RUNG
   // the same network as SCL:
   "Z256".ST_xSelectionManualMode := NOT "Z256".ST_xSelectionAutoMode;
END_REGION

REGION Network 12: Condition ok for manual mode
   RUNG wire#powerrail
      Contact( "AlwaysTRUE" )
      Coil( "Z256".ST_xConditionOKManualMode )
   END_RUNG
   // the same network as SCL:
   "Z256".ST_xConditionOKManualMode := "AlwaysTRUE";
END_REGION

